(* Logix 5000 project; controller MV vendor 1 type 14 code 217 rev 31.11; software revision 31.00; part 21 of 53 *)
(* tags used below, declared in another part *)
   CheckTimeMask : INT;
   CWD : CHECKWORD_FLAGS;
   Delphi_Does_Eng_Func : BOOL;
   MC_CH2_DR1 : PlantItem;   // CH2_DR1
   MC_CH2_DR2 : PlantItem;   // CH2_DR2
   MC_CH2_DRAIN : PlantItem;   // CH2_DRAIN
   MC_CH2_DT1 : PlantItem;   // CH2_DT1
   MC_CH2_DT2 : PlantItem;   // CH2_DT2
   MC_CH2_LF1 : PlantItem;   // CH2_LF1
   MC_CH2_PR1 : PlantItem;   // CH2_PR1
   MC_CH2_R2R : PlantItem;   // CH2_R2R
   MC_CH2_R3R : PlantItem;   // CH2_R3R
   MC_CH2_R4R : PlantItem;   // CH2_R4R
   MC_CH2_R5R : PlantItem;   // CH2_R5R
   MC_CH2_R6R : PlantItem;   // CH2_R6R
   MC_CH2_RR : PlantItem;   // CH2_RR
   MC_N255 : INT[255];   // CHECKWORDS Plant item checkword s
   TempChecktime : DINT;
(* MC_Common, continued *)

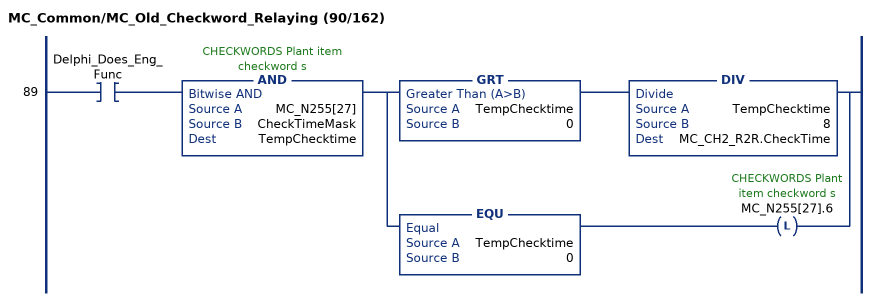
   [picture p361: MC_Common/MC_Old_Checkword_Relaying rungs 89-89]
   89: XIC(Delphi_Does_Eng_Func)AND(MC_N255[27],CheckTimeMask,TempChecktime)[GRT(TempChecktime,0) DIV(TempChecktime,8,MC_CH2_R2R.CheckTime) ,EQU(TempChecktime,0) OTL(MC_N255[27].6) ];
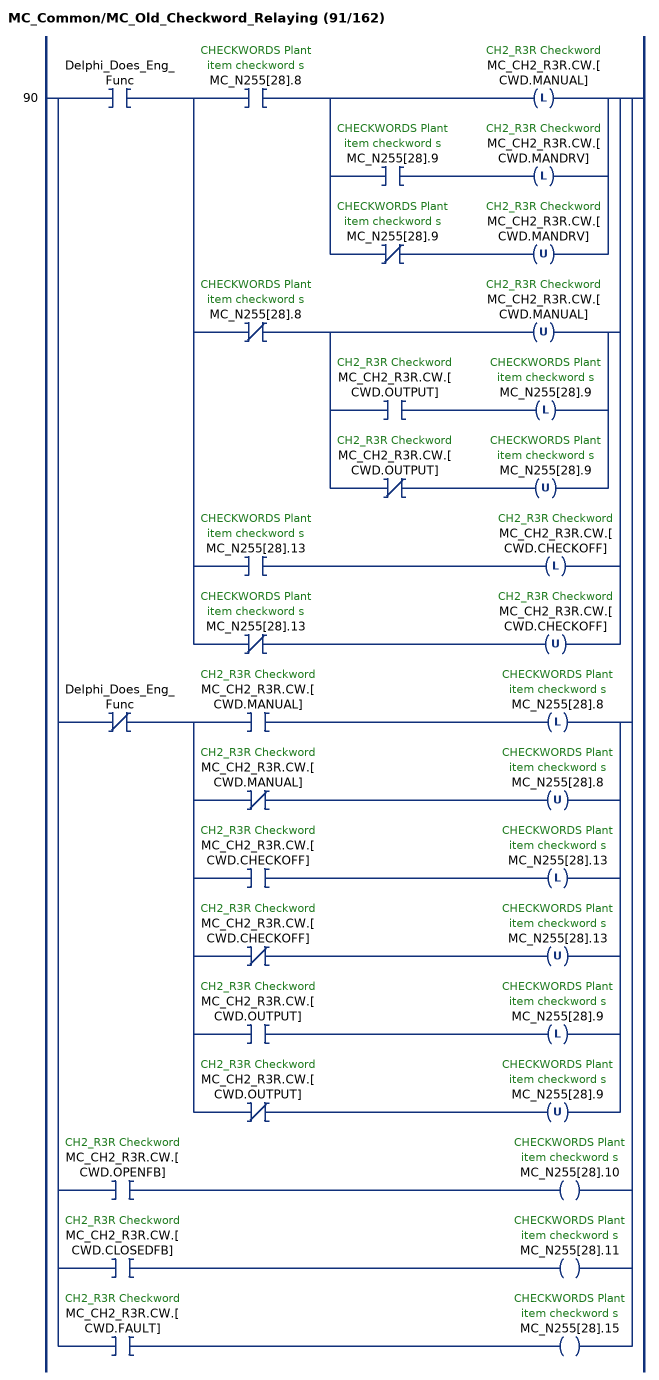
   90: [XIC(Delphi_Does_Eng_Func) [[XIC(MC_N255[28].8) [OTL(MC_CH2_R3R.CW.[CWD.MANUAL]) ,XIC(MC_N255[28].9) OTL(MC_CH2_R3R.CW.[CWD.MANDRV]) ,XIO(MC_N255[28].9) OTU(MC_CH2_R3R.CW.[CWD.MANDRV]) ] ,XIO(MC_N255[28].8) [OTU(MC_CH2_R3R.CW.[CWD.MANUAL]) ,[XIC(MC_CH2_R3R.CW.[CWD.OUTPUT]) OTL(MC_N255[28].9) ,XIO(MC_CH2_R3R.CW.[CWD.OUTPUT]) OTU(MC_N255[28].9) ] ] ] ,[XIC(MC_N255[28].13) OTL(MC_CH2_R3R.CW.[CWD.CHECKOFF]) ,XIO(MC_N255[28].13) OTU(MC_CH2_R3R.CW.[CWD.CHECKOFF]) ] ] ,XIO(Delphi_Does_Eng_Func) [[XIC(MC_CH2_R3R.CW.[CWD.MANUAL]) OTL(MC_N255[28].8) ,XIO(MC_CH2_R3R.CW.[CWD.MANUAL]) OTU(MC_N255[28].8) ] ,[XIC(MC_CH2_R3R.CW.[CWD.CHECKOFF]) OTL(MC_N255[28].13) ,XIO(MC_CH2_R3R.CW.[CWD.CHECKOFF]) OTU(MC_N255[28].13) ] ,[XIC(MC_CH2_R3R.CW.[CWD.OUTPUT]) OTL(MC_N255[28].9) ,XIO(MC_CH2_R3R.CW.[CWD.OUTPUT]) OTU(MC_N255[28].9) ] ] ,XIC(MC_CH2_R3R.CW.[CWD.OPENFB]) OTE(MC_N255[28].10) ,XIC(MC_CH2_R3R.CW.[CWD.CLOSEDFB]) OTE(MC_N255[28].11) ,XIC(MC_CH2_R3R.CW.[CWD.FAULT]) OTE(MC_N255[28].15) ];
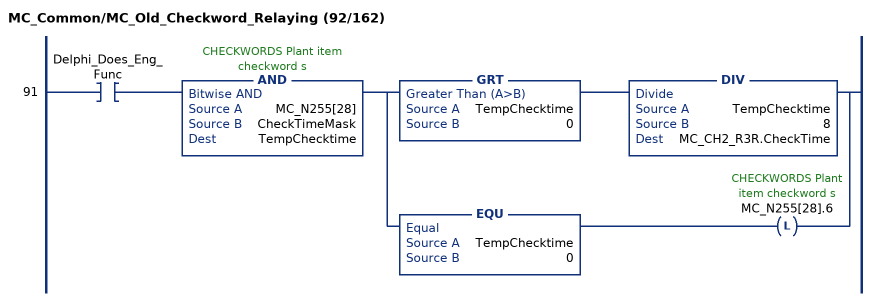
   91: XIC(Delphi_Does_Eng_Func)AND(MC_N255[28],CheckTimeMask,TempChecktime)[GRT(TempChecktime,0) DIV(TempChecktime,8,MC_CH2_R3R.CheckTime) ,EQU(TempChecktime,0) OTL(MC_N255[28].6) ];
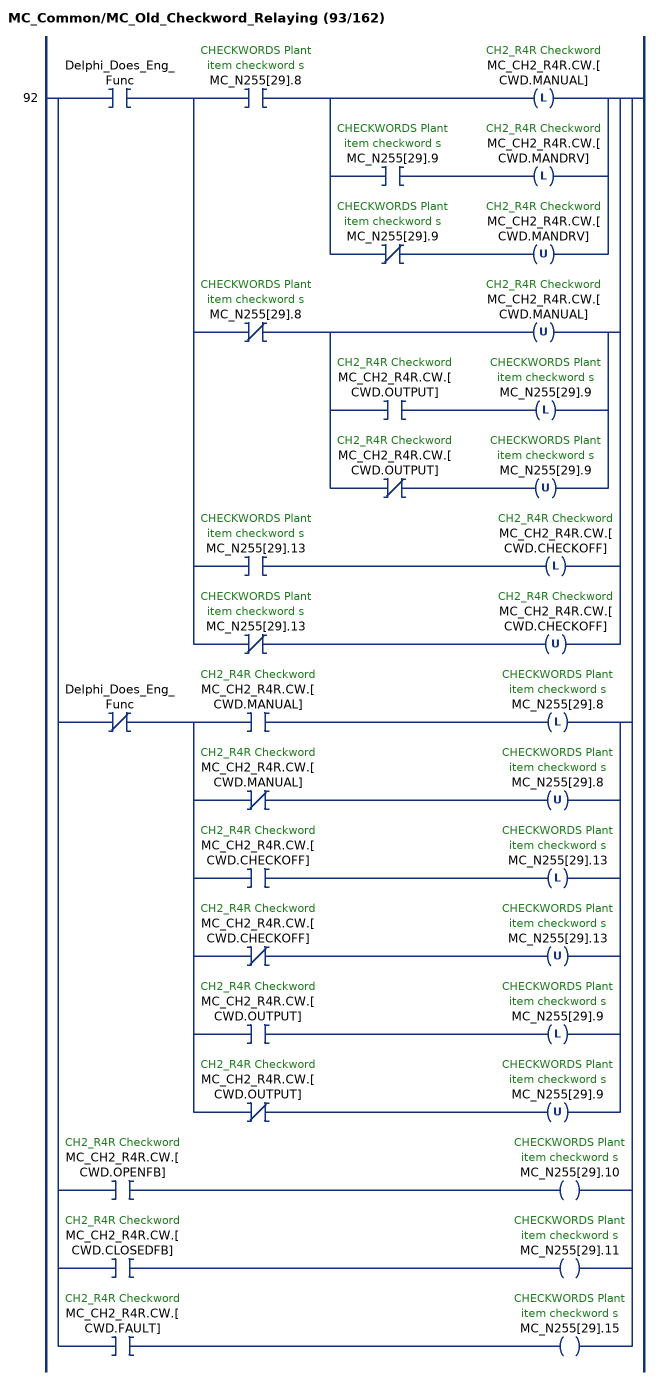
   92: [XIC(Delphi_Does_Eng_Func) [[XIC(MC_N255[29].8) [OTL(MC_CH2_R4R.CW.[CWD.MANUAL]) ,XIC(MC_N255[29].9) OTL(MC_CH2_R4R.CW.[CWD.MANDRV]) ,XIO(MC_N255[29].9) OTU(MC_CH2_R4R.CW.[CWD.MANDRV]) ] ,XIO(MC_N255[29].8) [OTU(MC_CH2_R4R.CW.[CWD.MANUAL]) ,[XIC(MC_CH2_R4R.CW.[CWD.OUTPUT]) OTL(MC_N255[29].9) ,XIO(MC_CH2_R4R.CW.[CWD.OUTPUT]) OTU(MC_N255[29].9) ] ] ] ,[XIC(MC_N255[29].13) OTL(MC_CH2_R4R.CW.[CWD.CHECKOFF]) ,XIO(MC_N255[29].13) OTU(MC_CH2_R4R.CW.[CWD.CHECKOFF]) ] ] ,XIO(Delphi_Does_Eng_Func) [[XIC(MC_CH2_R4R.CW.[CWD.MANUAL]) OTL(MC_N255[29].8) ,XIO(MC_CH2_R4R.CW.[CWD.MANUAL]) OTU(MC_N255[29].8) ] ,[XIC(MC_CH2_R4R.CW.[CWD.CHECKOFF]) OTL(MC_N255[29].13) ,XIO(MC_CH2_R4R.CW.[CWD.CHECKOFF]) OTU(MC_N255[29].13) ] ,[XIC(MC_CH2_R4R.CW.[CWD.OUTPUT]) OTL(MC_N255[29].9) ,XIO(MC_CH2_R4R.CW.[CWD.OUTPUT]) OTU(MC_N255[29].9) ] ] ,XIC(MC_CH2_R4R.CW.[CWD.OPENFB]) OTE(MC_N255[29].10) ,XIC(MC_CH2_R4R.CW.[CWD.CLOSEDFB]) OTE(MC_N255[29].11) ,XIC(MC_CH2_R4R.CW.[CWD.FAULT]) OTE(MC_N255[29].15) ];
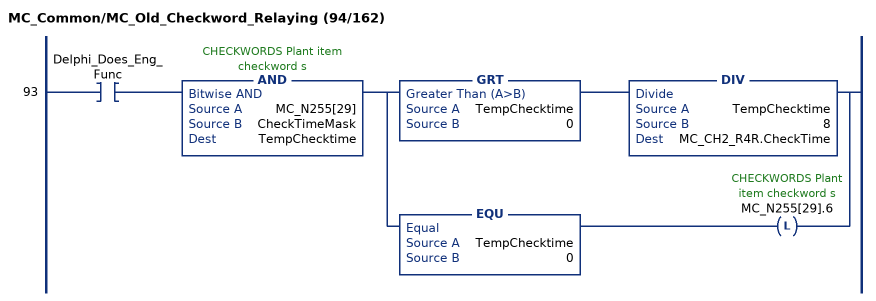
   93: XIC(Delphi_Does_Eng_Func)AND(MC_N255[29],CheckTimeMask,TempChecktime)[GRT(TempChecktime,0) DIV(TempChecktime,8,MC_CH2_R4R.CheckTime) ,EQU(TempChecktime,0) OTL(MC_N255[29].6) ];
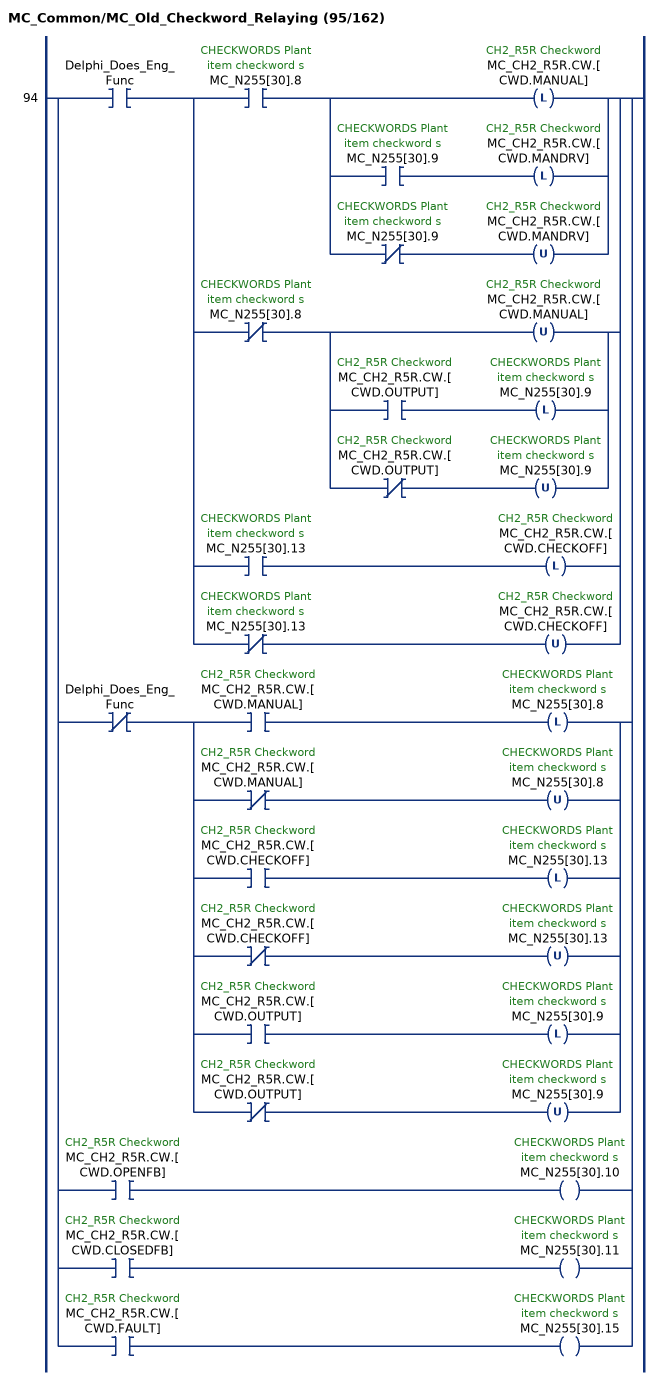
   94: [XIC(Delphi_Does_Eng_Func) [[XIC(MC_N255[30].8) [OTL(MC_CH2_R5R.CW.[CWD.MANUAL]) ,XIC(MC_N255[30].9) OTL(MC_CH2_R5R.CW.[CWD.MANDRV]) ,XIO(MC_N255[30].9) OTU(MC_CH2_R5R.CW.[CWD.MANDRV]) ] ,XIO(MC_N255[30].8) [OTU(MC_CH2_R5R.CW.[CWD.MANUAL]) ,[XIC(MC_CH2_R5R.CW.[CWD.OUTPUT]) OTL(MC_N255[30].9) ,XIO(MC_CH2_R5R.CW.[CWD.OUTPUT]) OTU(MC_N255[30].9) ] ] ] ,[XIC(MC_N255[30].13) OTL(MC_CH2_R5R.CW.[CWD.CHECKOFF]) ,XIO(MC_N255[30].13) OTU(MC_CH2_R5R.CW.[CWD.CHECKOFF]) ] ] ,XIO(Delphi_Does_Eng_Func) [[XIC(MC_CH2_R5R.CW.[CWD.MANUAL]) OTL(MC_N255[30].8) ,XIO(MC_CH2_R5R.CW.[CWD.MANUAL]) OTU(MC_N255[30].8) ] ,[XIC(MC_CH2_R5R.CW.[CWD.CHECKOFF]) OTL(MC_N255[30].13) ,XIO(MC_CH2_R5R.CW.[CWD.CHECKOFF]) OTU(MC_N255[30].13) ] ,[XIC(MC_CH2_R5R.CW.[CWD.OUTPUT]) OTL(MC_N255[30].9) ,XIO(MC_CH2_R5R.CW.[CWD.OUTPUT]) OTU(MC_N255[30].9) ] ] ,XIC(MC_CH2_R5R.CW.[CWD.OPENFB]) OTE(MC_N255[30].10) ,XIC(MC_CH2_R5R.CW.[CWD.CLOSEDFB]) OTE(MC_N255[30].11) ,XIC(MC_CH2_R5R.CW.[CWD.FAULT]) OTE(MC_N255[30].15) ];
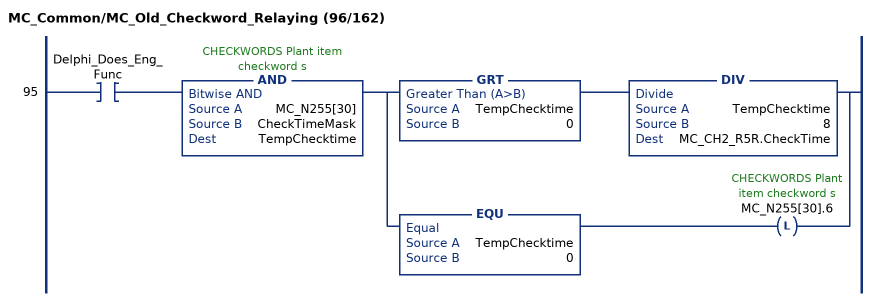
   95: XIC(Delphi_Does_Eng_Func)AND(MC_N255[30],CheckTimeMask,TempChecktime)[GRT(TempChecktime,0) DIV(TempChecktime,8,MC_CH2_R5R.CheckTime) ,EQU(TempChecktime,0) OTL(MC_N255[30].6) ];
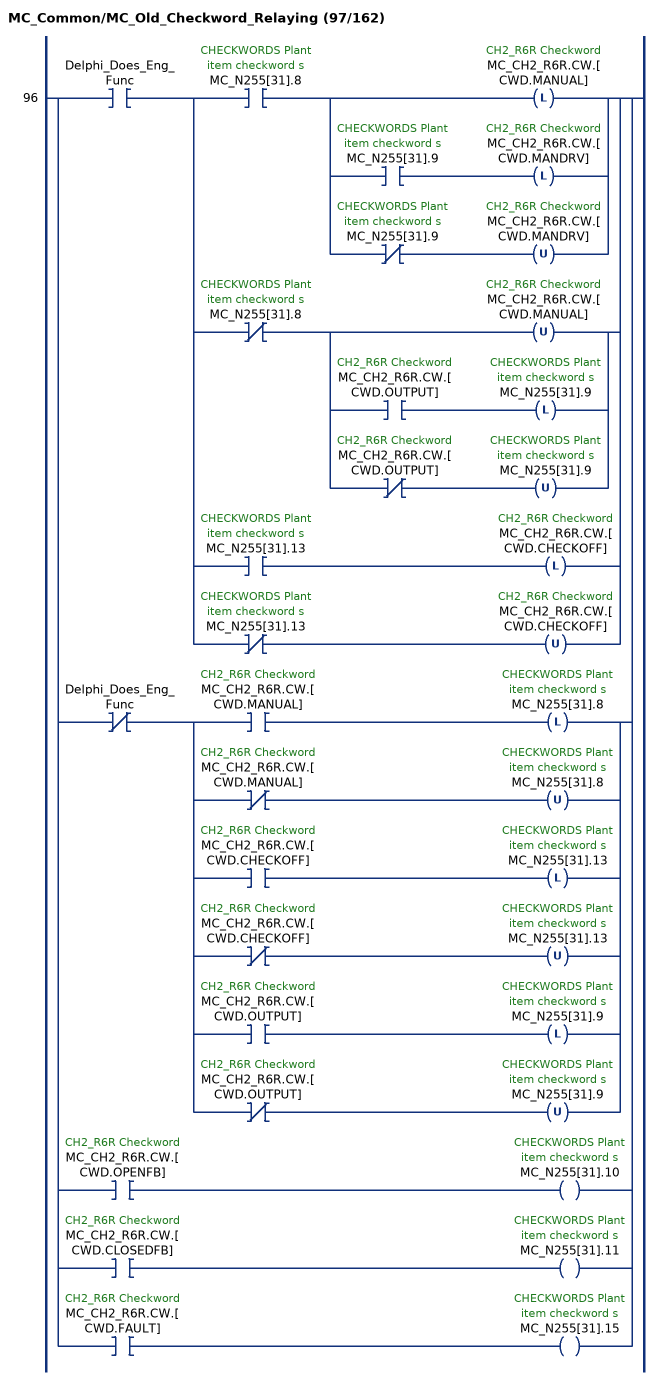
   96: [XIC(Delphi_Does_Eng_Func) [[XIC(MC_N255[31].8) [OTL(MC_CH2_R6R.CW.[CWD.MANUAL]) ,XIC(MC_N255[31].9) OTL(MC_CH2_R6R.CW.[CWD.MANDRV]) ,XIO(MC_N255[31].9) OTU(MC_CH2_R6R.CW.[CWD.MANDRV]) ] ,XIO(MC_N255[31].8) [OTU(MC_CH2_R6R.CW.[CWD.MANUAL]) ,[XIC(MC_CH2_R6R.CW.[CWD.OUTPUT]) OTL(MC_N255[31].9) ,XIO(MC_CH2_R6R.CW.[CWD.OUTPUT]) OTU(MC_N255[31].9) ] ] ] ,[XIC(MC_N255[31].13) OTL(MC_CH2_R6R.CW.[CWD.CHECKOFF]) ,XIO(MC_N255[31].13) OTU(MC_CH2_R6R.CW.[CWD.CHECKOFF]) ] ] ,XIO(Delphi_Does_Eng_Func) [[XIC(MC_CH2_R6R.CW.[CWD.MANUAL]) OTL(MC_N255[31].8) ,XIO(MC_CH2_R6R.CW.[CWD.MANUAL]) OTU(MC_N255[31].8) ] ,[XIC(MC_CH2_R6R.CW.[CWD.CHECKOFF]) OTL(MC_N255[31].13) ,XIO(MC_CH2_R6R.CW.[CWD.CHECKOFF]) OTU(MC_N255[31].13) ] ,[XIC(MC_CH2_R6R.CW.[CWD.OUTPUT]) OTL(MC_N255[31].9) ,XIO(MC_CH2_R6R.CW.[CWD.OUTPUT]) OTU(MC_N255[31].9) ] ] ,XIC(MC_CH2_R6R.CW.[CWD.OPENFB]) OTE(MC_N255[31].10) ,XIC(MC_CH2_R6R.CW.[CWD.CLOSEDFB]) OTE(MC_N255[31].11) ,XIC(MC_CH2_R6R.CW.[CWD.FAULT]) OTE(MC_N255[31].15) ];
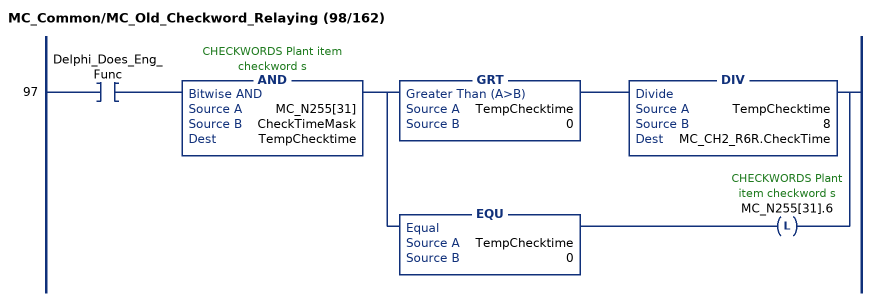
   97: XIC(Delphi_Does_Eng_Func)AND(MC_N255[31],CheckTimeMask,TempChecktime)[GRT(TempChecktime,0) DIV(TempChecktime,8,MC_CH2_R6R.CheckTime) ,EQU(TempChecktime,0) OTL(MC_N255[31].6) ];
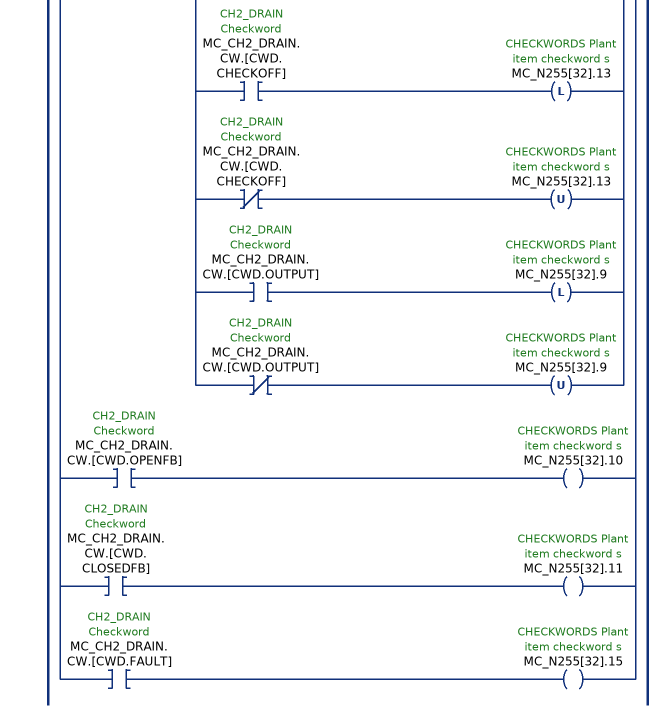
   98: [XIC(Delphi_Does_Eng_Func) [[XIC(MC_N255[32].8) [OTL(MC_CH2_DRAIN.CW.[CWD.MANUAL]) ,XIC(MC_N255[32].9) OTL(MC_CH2_DRAIN.CW.[CWD.MANDRV]) ,XIO(MC_N255[32].9) OTU(MC_CH2_DRAIN.CW.[CWD.MANDRV]) ] ,XIO(MC_N255[32].8) [OTU(MC_CH2_DRAIN.CW.[CWD.MANUAL]) ,[XIC(MC_CH2_DRAIN.CW.[CWD.OUTPUT]) OTL(MC_N255[32].9) ,XIO(MC_CH2_DRAIN.CW.[CWD.OUTPUT]) OTU(MC_N255[32].9) ] ] ] ,[XIC(MC_N255[32].13) OTL(MC_CH2_DRAIN.CW.[CWD.CHECKOFF]) ,XIO(MC_N255[32].13) OTU(MC_CH2_DRAIN.CW.[CWD.CHECKOFF]) ] ] ,XIO(Delphi_Does_Eng_Func) [[XIC(MC_CH2_DRAIN.CW.[CWD.MANUAL]) OTL(MC_N255[32].8) ,XIO(MC_CH2_DRAIN.CW.[CWD.MANUAL]) OTU(MC_N255[32].8) ] ,[XIC(MC_CH2_DRAIN.CW.[CWD.CHECKOFF]) OTL(MC_N255[32].13) ,XIO(MC_CH2_DRAIN.CW.[CWD.CHECKOFF]) OTU(MC_N255[32].13) ] ,[XIC(MC_CH2_DRAIN.CW.[CWD.OUTPUT]) OTL(MC_N255[32].9) ,XIO(MC_CH2_DRAIN.CW.[CWD.OUTPUT]) OTU(MC_N255[32].9) ] ] ,XIC(MC_CH2_DRAIN.CW.[CWD.OPENFB]) OTE(MC_N255[32].10) ,XIC(MC_CH2_DRAIN.CW.[CWD.CLOSEDFB]) OTE(MC_N255[32].11) ,XIC(MC_CH2_DRAIN.CW.[CWD.FAULT]) OTE(MC_N255[32].15) ];
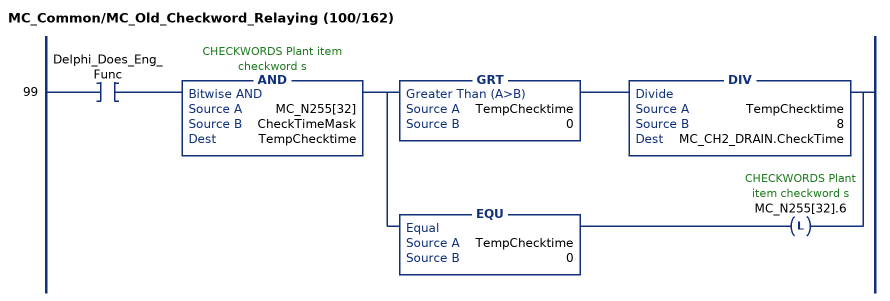
   99: XIC(Delphi_Does_Eng_Func)AND(MC_N255[32],CheckTimeMask,TempChecktime)[GRT(TempChecktime,0) DIV(TempChecktime,8,MC_CH2_DRAIN.CheckTime) ,EQU(TempChecktime,0) OTL(MC_N255[32].6) ];
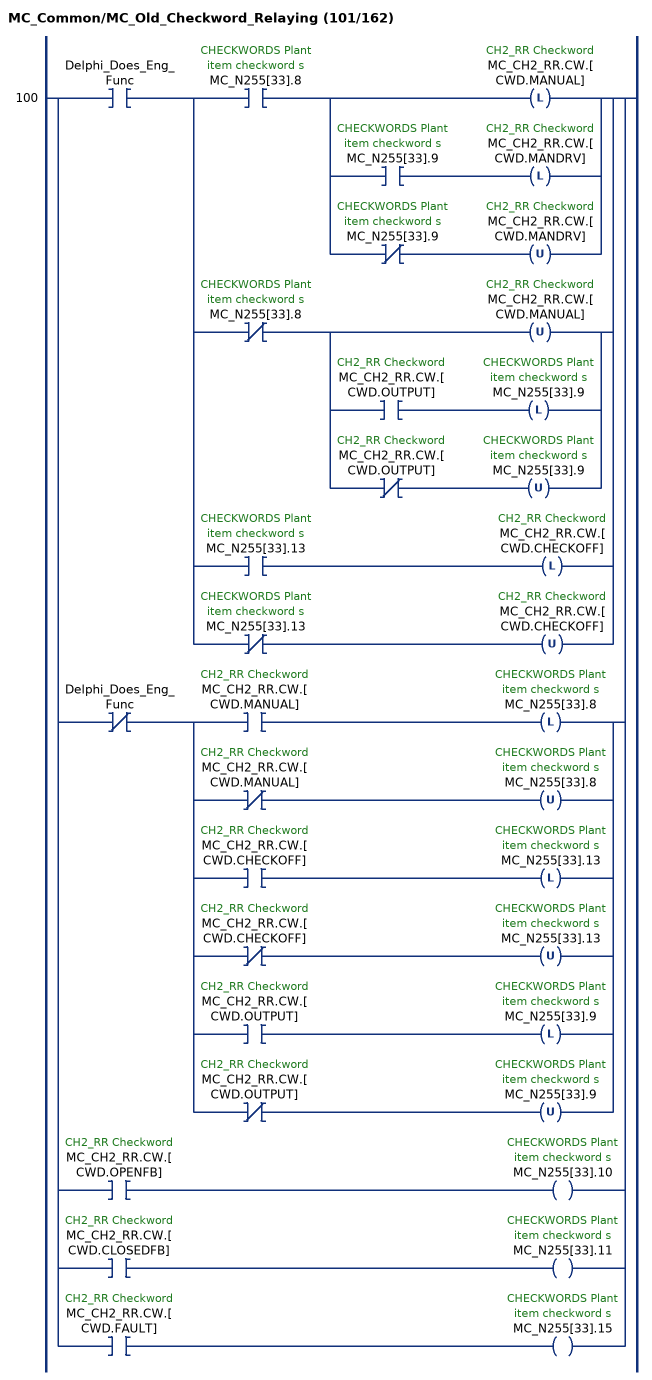
   100: [XIC(Delphi_Does_Eng_Func) [[XIC(MC_N255[33].8) [OTL(MC_CH2_RR.CW.[CWD.MANUAL]) ,XIC(MC_N255[33].9) OTL(MC_CH2_RR.CW.[CWD.MANDRV]) ,XIO(MC_N255[33].9) OTU(MC_CH2_RR.CW.[CWD.MANDRV]) ] ,XIO(MC_N255[33].8) [OTU(MC_CH2_RR.CW.[CWD.MANUAL]) ,[XIC(MC_CH2_RR.CW.[CWD.OUTPUT]) OTL(MC_N255[33].9) ,XIO(MC_CH2_RR.CW.[CWD.OUTPUT]) OTU(MC_N255[33].9) ] ] ] ,[XIC(MC_N255[33].13) OTL(MC_CH2_RR.CW.[CWD.CHECKOFF]) ,XIO(MC_N255[33].13) OTU(MC_CH2_RR.CW.[CWD.CHECKOFF]) ] ] ,XIO(Delphi_Does_Eng_Func) [[XIC(MC_CH2_RR.CW.[CWD.MANUAL]) OTL(MC_N255[33].8) ,XIO(MC_CH2_RR.CW.[CWD.MANUAL]) OTU(MC_N255[33].8) ] ,[XIC(MC_CH2_RR.CW.[CWD.CHECKOFF]) OTL(MC_N255[33].13) ,XIO(MC_CH2_RR.CW.[CWD.CHECKOFF]) OTU(MC_N255[33].13) ] ,[XIC(MC_CH2_RR.CW.[CWD.OUTPUT]) OTL(MC_N255[33].9) ,XIO(MC_CH2_RR.CW.[CWD.OUTPUT]) OTU(MC_N255[33].9) ] ] ,XIC(MC_CH2_RR.CW.[CWD.OPENFB]) OTE(MC_N255[33].10) ,XIC(MC_CH2_RR.CW.[CWD.CLOSEDFB]) OTE(MC_N255[33].11) ,XIC(MC_CH2_RR.CW.[CWD.FAULT]) OTE(MC_N255[33].15) ];
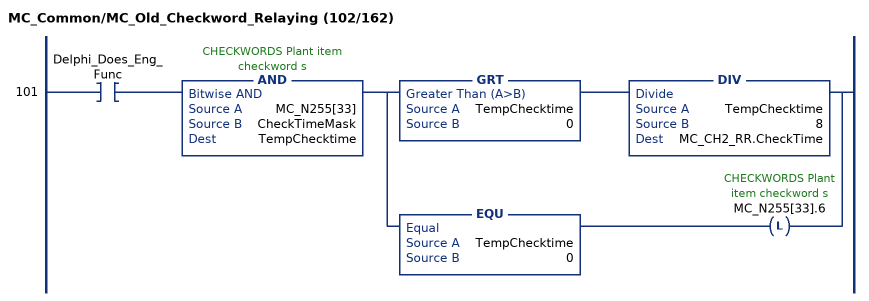
   101: XIC(Delphi_Does_Eng_Func)AND(MC_N255[33],CheckTimeMask,TempChecktime)[GRT(TempChecktime,0) DIV(TempChecktime,8,MC_CH2_RR.CheckTime) ,EQU(TempChecktime,0) OTL(MC_N255[33].6) ];
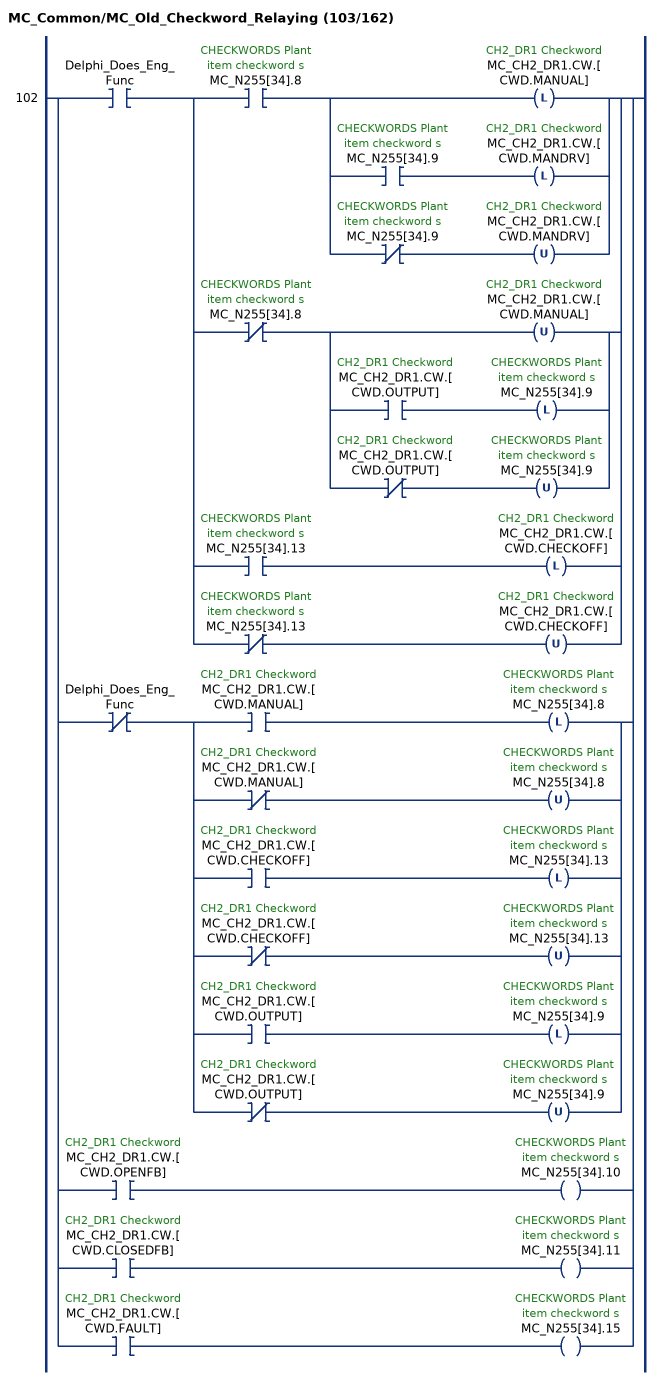
   102: [XIC(Delphi_Does_Eng_Func) [[XIC(MC_N255[34].8) [OTL(MC_CH2_DR1.CW.[CWD.MANUAL]) ,XIC(MC_N255[34].9) OTL(MC_CH2_DR1.CW.[CWD.MANDRV]) ,XIO(MC_N255[34].9) OTU(MC_CH2_DR1.CW.[CWD.MANDRV]) ] ,XIO(MC_N255[34].8) [OTU(MC_CH2_DR1.CW.[CWD.MANUAL]) ,[XIC(MC_CH2_DR1.CW.[CWD.OUTPUT]) OTL(MC_N255[34].9) ,XIO(MC_CH2_DR1.CW.[CWD.OUTPUT]) OTU(MC_N255[34].9) ] ] ] ,[XIC(MC_N255[34].13) OTL(MC_CH2_DR1.CW.[CWD.CHECKOFF]) ,XIO(MC_N255[34].13) OTU(MC_CH2_DR1.CW.[CWD.CHECKOFF]) ] ] ,XIO(Delphi_Does_Eng_Func) [[XIC(MC_CH2_DR1.CW.[CWD.MANUAL]) OTL(MC_N255[34].8) ,XIO(MC_CH2_DR1.CW.[CWD.MANUAL]) OTU(MC_N255[34].8) ] ,[XIC(MC_CH2_DR1.CW.[CWD.CHECKOFF]) OTL(MC_N255[34].13) ,XIO(MC_CH2_DR1.CW.[CWD.CHECKOFF]) OTU(MC_N255[34].13) ] ,[XIC(MC_CH2_DR1.CW.[CWD.OUTPUT]) OTL(MC_N255[34].9) ,XIO(MC_CH2_DR1.CW.[CWD.OUTPUT]) OTU(MC_N255[34].9) ] ] ,XIC(MC_CH2_DR1.CW.[CWD.OPENFB]) OTE(MC_N255[34].10) ,XIC(MC_CH2_DR1.CW.[CWD.CLOSEDFB]) OTE(MC_N255[34].11) ,XIC(MC_CH2_DR1.CW.[CWD.FAULT]) OTE(MC_N255[34].15) ];
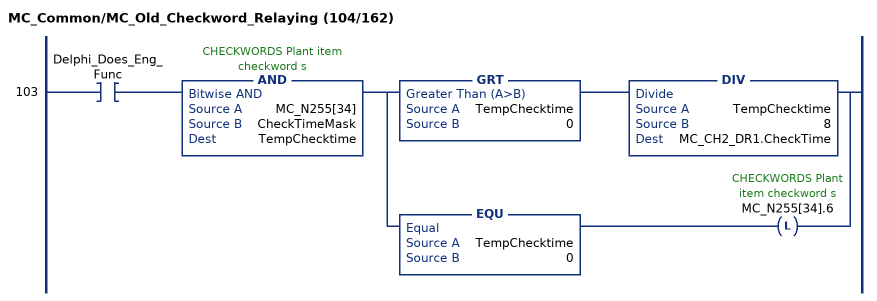
   103: XIC(Delphi_Does_Eng_Func)AND(MC_N255[34],CheckTimeMask,TempChecktime)[GRT(TempChecktime,0) DIV(TempChecktime,8,MC_CH2_DR1.CheckTime) ,EQU(TempChecktime,0) OTL(MC_N255[34].6) ];
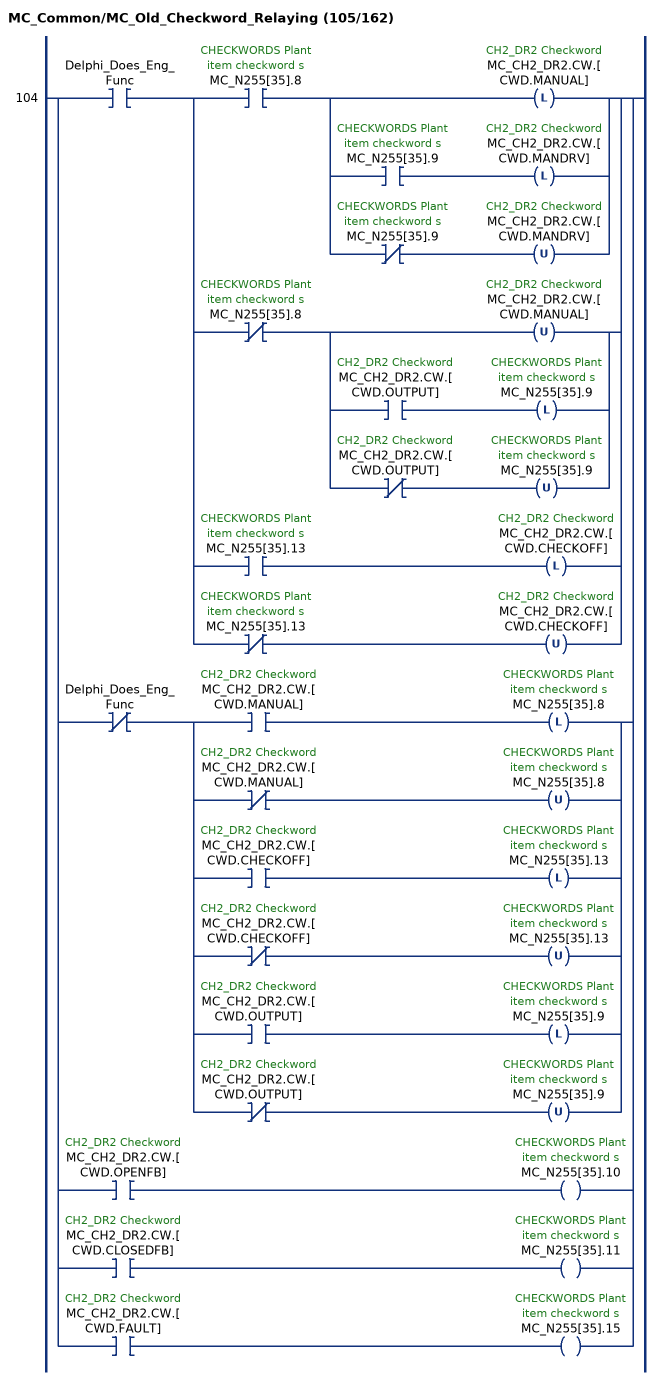
   104: [XIC(Delphi_Does_Eng_Func) [[XIC(MC_N255[35].8) [OTL(MC_CH2_DR2.CW.[CWD.MANUAL]) ,XIC(MC_N255[35].9) OTL(MC_CH2_DR2.CW.[CWD.MANDRV]) ,XIO(MC_N255[35].9) OTU(MC_CH2_DR2.CW.[CWD.MANDRV]) ] ,XIO(MC_N255[35].8) [OTU(MC_CH2_DR2.CW.[CWD.MANUAL]) ,[XIC(MC_CH2_DR2.CW.[CWD.OUTPUT]) OTL(MC_N255[35].9) ,XIO(MC_CH2_DR2.CW.[CWD.OUTPUT]) OTU(MC_N255[35].9) ] ] ] ,[XIC(MC_N255[35].13) OTL(MC_CH2_DR2.CW.[CWD.CHECKOFF]) ,XIO(MC_N255[35].13) OTU(MC_CH2_DR2.CW.[CWD.CHECKOFF]) ] ] ,XIO(Delphi_Does_Eng_Func) [[XIC(MC_CH2_DR2.CW.[CWD.MANUAL]) OTL(MC_N255[35].8) ,XIO(MC_CH2_DR2.CW.[CWD.MANUAL]) OTU(MC_N255[35].8) ] ,[XIC(MC_CH2_DR2.CW.[CWD.CHECKOFF]) OTL(MC_N255[35].13) ,XIO(MC_CH2_DR2.CW.[CWD.CHECKOFF]) OTU(MC_N255[35].13) ] ,[XIC(MC_CH2_DR2.CW.[CWD.OUTPUT]) OTL(MC_N255[35].9) ,XIO(MC_CH2_DR2.CW.[CWD.OUTPUT]) OTU(MC_N255[35].9) ] ] ,XIC(MC_CH2_DR2.CW.[CWD.OPENFB]) OTE(MC_N255[35].10) ,XIC(MC_CH2_DR2.CW.[CWD.CLOSEDFB]) OTE(MC_N255[35].11) ,XIC(MC_CH2_DR2.CW.[CWD.FAULT]) OTE(MC_N255[35].15) ];
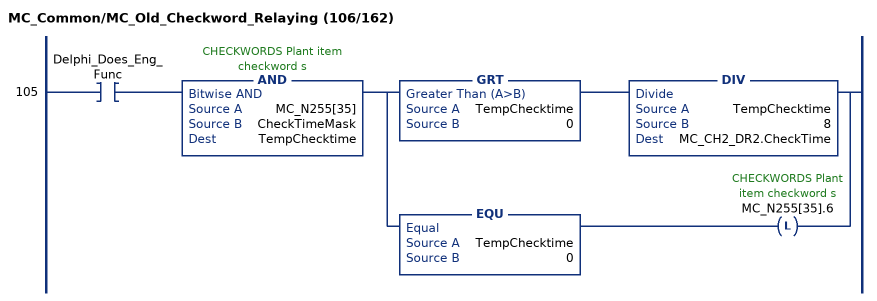
   105: XIC(Delphi_Does_Eng_Func)AND(MC_N255[35],CheckTimeMask,TempChecktime)[GRT(TempChecktime,0) DIV(TempChecktime,8,MC_CH2_DR2.CheckTime) ,EQU(TempChecktime,0) OTL(MC_N255[35].6) ];
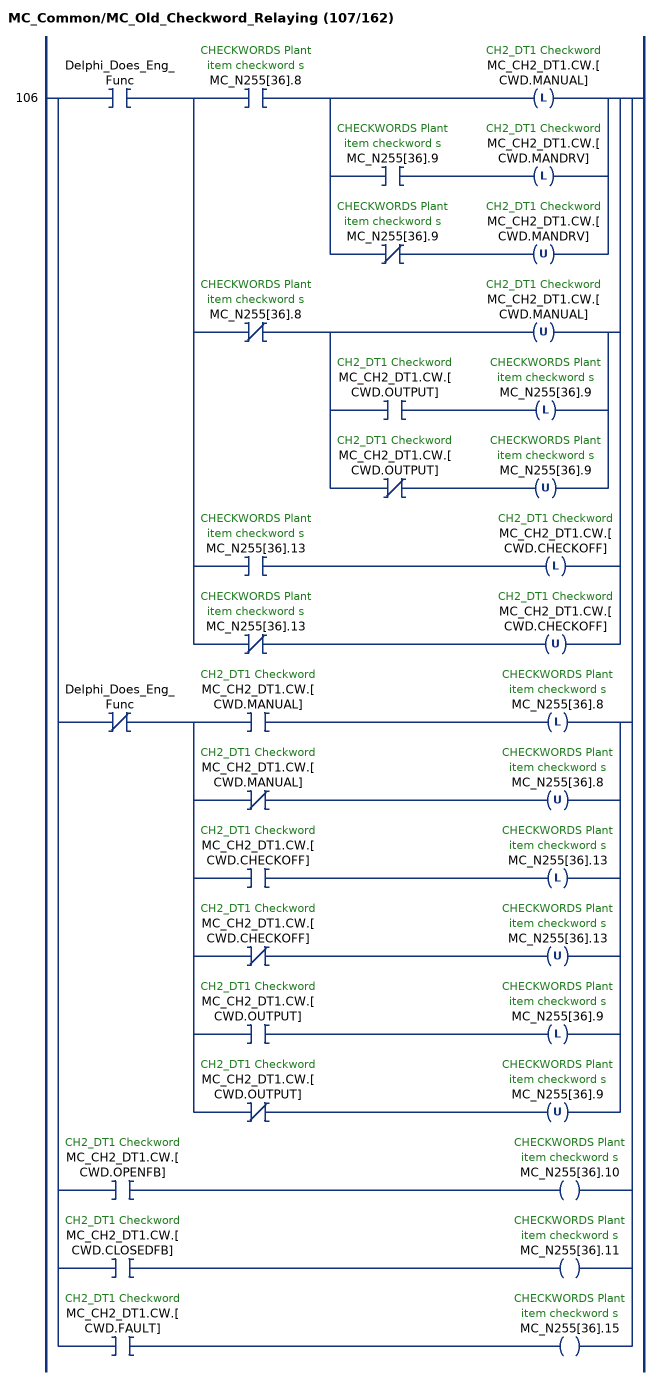
   106: [XIC(Delphi_Does_Eng_Func) [[XIC(MC_N255[36].8) [OTL(MC_CH2_DT1.CW.[CWD.MANUAL]) ,XIC(MC_N255[36].9) OTL(MC_CH2_DT1.CW.[CWD.MANDRV]) ,XIO(MC_N255[36].9) OTU(MC_CH2_DT1.CW.[CWD.MANDRV]) ] ,XIO(MC_N255[36].8) [OTU(MC_CH2_DT1.CW.[CWD.MANUAL]) ,[XIC(MC_CH2_DT1.CW.[CWD.OUTPUT]) OTL(MC_N255[36].9) ,XIO(MC_CH2_DT1.CW.[CWD.OUTPUT]) OTU(MC_N255[36].9) ] ] ] ,[XIC(MC_N255[36].13) OTL(MC_CH2_DT1.CW.[CWD.CHECKOFF]) ,XIO(MC_N255[36].13) OTU(MC_CH2_DT1.CW.[CWD.CHECKOFF]) ] ] ,XIO(Delphi_Does_Eng_Func) [[XIC(MC_CH2_DT1.CW.[CWD.MANUAL]) OTL(MC_N255[36].8) ,XIO(MC_CH2_DT1.CW.[CWD.MANUAL]) OTU(MC_N255[36].8) ] ,[XIC(MC_CH2_DT1.CW.[CWD.CHECKOFF]) OTL(MC_N255[36].13) ,XIO(MC_CH2_DT1.CW.[CWD.CHECKOFF]) OTU(MC_N255[36].13) ] ,[XIC(MC_CH2_DT1.CW.[CWD.OUTPUT]) OTL(MC_N255[36].9) ,XIO(MC_CH2_DT1.CW.[CWD.OUTPUT]) OTU(MC_N255[36].9) ] ] ,XIC(MC_CH2_DT1.CW.[CWD.OPENFB]) OTE(MC_N255[36].10) ,XIC(MC_CH2_DT1.CW.[CWD.CLOSEDFB]) OTE(MC_N255[36].11) ,XIC(MC_CH2_DT1.CW.[CWD.FAULT]) OTE(MC_N255[36].15) ];
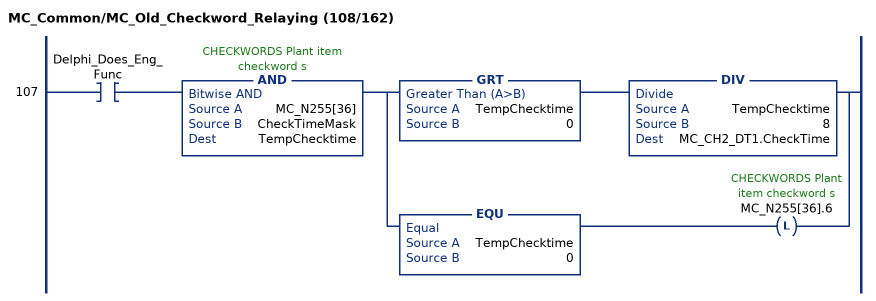
   107: XIC(Delphi_Does_Eng_Func)AND(MC_N255[36],CheckTimeMask,TempChecktime)[GRT(TempChecktime,0) DIV(TempChecktime,8,MC_CH2_DT1.CheckTime) ,EQU(TempChecktime,0) OTL(MC_N255[36].6) ];
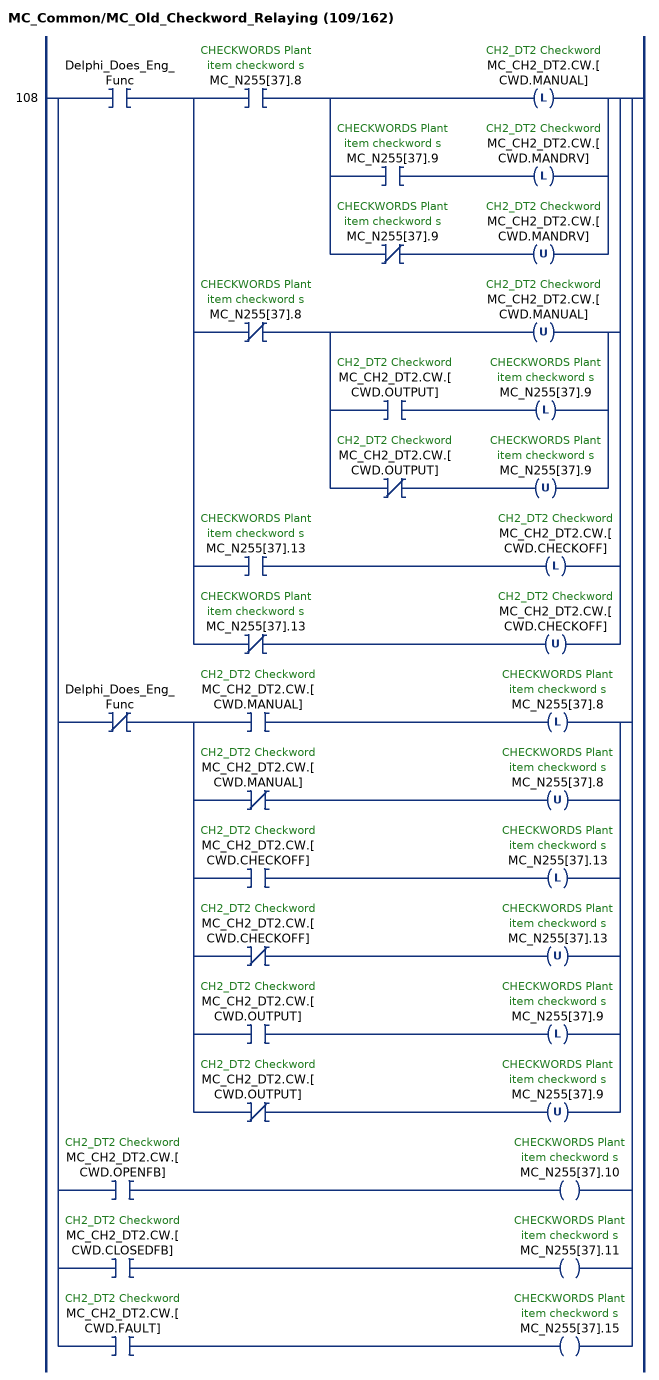
   108: [XIC(Delphi_Does_Eng_Func) [[XIC(MC_N255[37].8) [OTL(MC_CH2_DT2.CW.[CWD.MANUAL]) ,XIC(MC_N255[37].9) OTL(MC_CH2_DT2.CW.[CWD.MANDRV]) ,XIO(MC_N255[37].9) OTU(MC_CH2_DT2.CW.[CWD.MANDRV]) ] ,XIO(MC_N255[37].8) [OTU(MC_CH2_DT2.CW.[CWD.MANUAL]) ,[XIC(MC_CH2_DT2.CW.[CWD.OUTPUT]) OTL(MC_N255[37].9) ,XIO(MC_CH2_DT2.CW.[CWD.OUTPUT]) OTU(MC_N255[37].9) ] ] ] ,[XIC(MC_N255[37].13) OTL(MC_CH2_DT2.CW.[CWD.CHECKOFF]) ,XIO(MC_N255[37].13) OTU(MC_CH2_DT2.CW.[CWD.CHECKOFF]) ] ] ,XIO(Delphi_Does_Eng_Func) [[XIC(MC_CH2_DT2.CW.[CWD.MANUAL]) OTL(MC_N255[37].8) ,XIO(MC_CH2_DT2.CW.[CWD.MANUAL]) OTU(MC_N255[37].8) ] ,[XIC(MC_CH2_DT2.CW.[CWD.CHECKOFF]) OTL(MC_N255[37].13) ,XIO(MC_CH2_DT2.CW.[CWD.CHECKOFF]) OTU(MC_N255[37].13) ] ,[XIC(MC_CH2_DT2.CW.[CWD.OUTPUT]) OTL(MC_N255[37].9) ,XIO(MC_CH2_DT2.CW.[CWD.OUTPUT]) OTU(MC_N255[37].9) ] ] ,XIC(MC_CH2_DT2.CW.[CWD.OPENFB]) OTE(MC_N255[37].10) ,XIC(MC_CH2_DT2.CW.[CWD.CLOSEDFB]) OTE(MC_N255[37].11) ,XIC(MC_CH2_DT2.CW.[CWD.FAULT]) OTE(MC_N255[37].15) ];
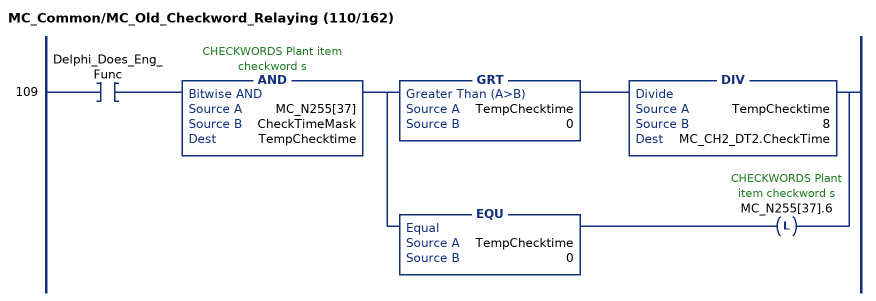
   109: XIC(Delphi_Does_Eng_Func)AND(MC_N255[37],CheckTimeMask,TempChecktime)[GRT(TempChecktime,0) DIV(TempChecktime,8,MC_CH2_DT2.CheckTime) ,EQU(TempChecktime,0) OTL(MC_N255[37].6) ];
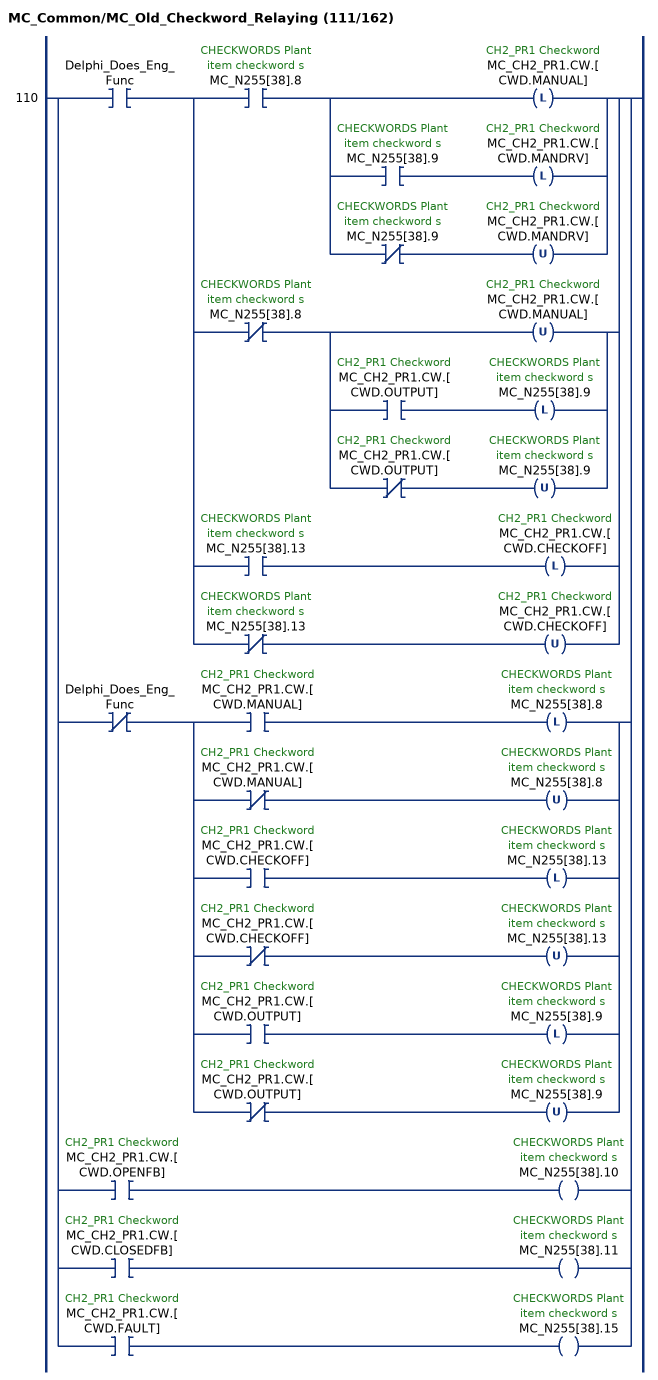
   110: [XIC(Delphi_Does_Eng_Func) [[XIC(MC_N255[38].8) [OTL(MC_CH2_PR1.CW.[CWD.MANUAL]) ,XIC(MC_N255[38].9) OTL(MC_CH2_PR1.CW.[CWD.MANDRV]) ,XIO(MC_N255[38].9) OTU(MC_CH2_PR1.CW.[CWD.MANDRV]) ] ,XIO(MC_N255[38].8) [OTU(MC_CH2_PR1.CW.[CWD.MANUAL]) ,[XIC(MC_CH2_PR1.CW.[CWD.OUTPUT]) OTL(MC_N255[38].9) ,XIO(MC_CH2_PR1.CW.[CWD.OUTPUT]) OTU(MC_N255[38].9) ] ] ] ,[XIC(MC_N255[38].13) OTL(MC_CH2_PR1.CW.[CWD.CHECKOFF]) ,XIO(MC_N255[38].13) OTU(MC_CH2_PR1.CW.[CWD.CHECKOFF]) ] ] ,XIO(Delphi_Does_Eng_Func) [[XIC(MC_CH2_PR1.CW.[CWD.MANUAL]) OTL(MC_N255[38].8) ,XIO(MC_CH2_PR1.CW.[CWD.MANUAL]) OTU(MC_N255[38].8) ] ,[XIC(MC_CH2_PR1.CW.[CWD.CHECKOFF]) OTL(MC_N255[38].13) ,XIO(MC_CH2_PR1.CW.[CWD.CHECKOFF]) OTU(MC_N255[38].13) ] ,[XIC(MC_CH2_PR1.CW.[CWD.OUTPUT]) OTL(MC_N255[38].9) ,XIO(MC_CH2_PR1.CW.[CWD.OUTPUT]) OTU(MC_N255[38].9) ] ] ,XIC(MC_CH2_PR1.CW.[CWD.OPENFB]) OTE(MC_N255[38].10) ,XIC(MC_CH2_PR1.CW.[CWD.CLOSEDFB]) OTE(MC_N255[38].11) ,XIC(MC_CH2_PR1.CW.[CWD.FAULT]) OTE(MC_N255[38].15) ];
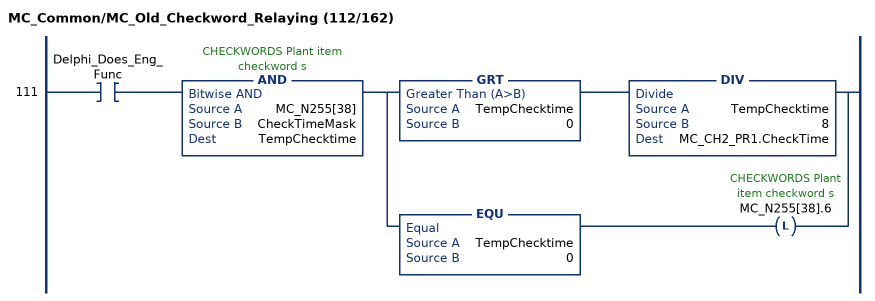
   111: XIC(Delphi_Does_Eng_Func)AND(MC_N255[38],CheckTimeMask,TempChecktime)[GRT(TempChecktime,0) DIV(TempChecktime,8,MC_CH2_PR1.CheckTime) ,EQU(TempChecktime,0) OTL(MC_N255[38].6) ];
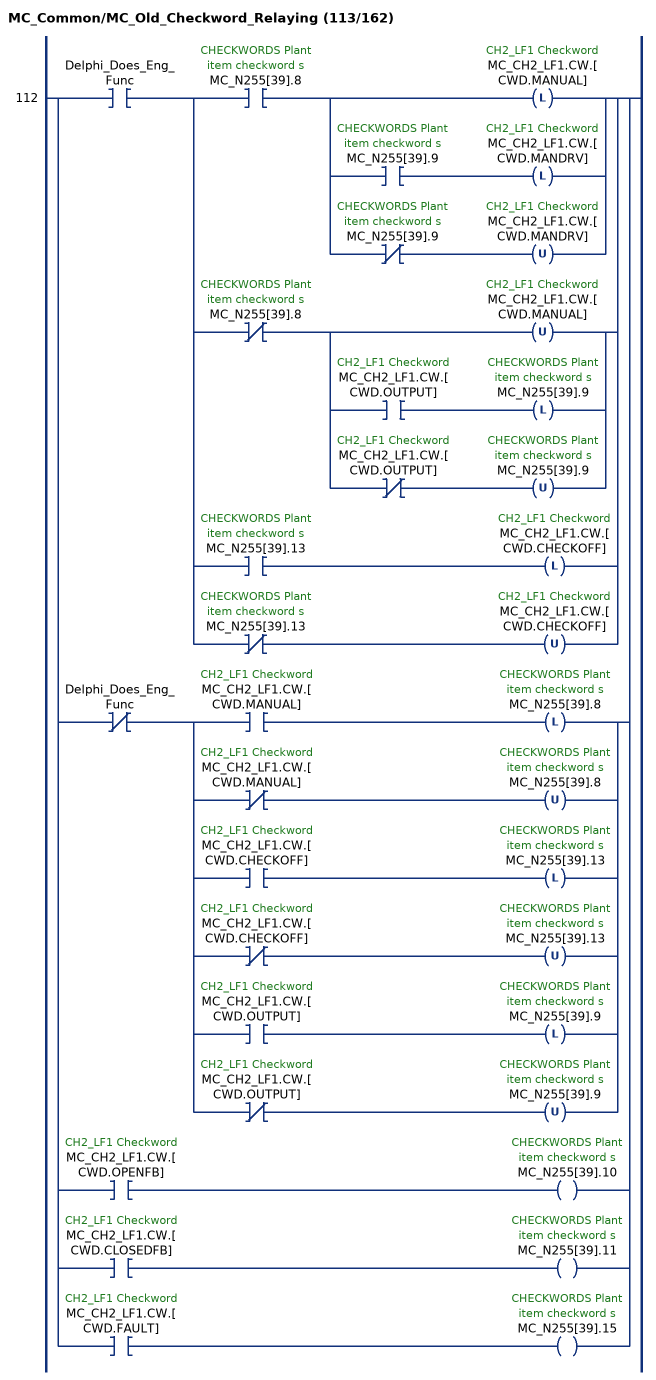
   112: [XIC(Delphi_Does_Eng_Func) [[XIC(MC_N255[39].8) [OTL(MC_CH2_LF1.CW.[CWD.MANUAL]) ,XIC(MC_N255[39].9) OTL(MC_CH2_LF1.CW.[CWD.MANDRV]) ,XIO(MC_N255[39].9) OTU(MC_CH2_LF1.CW.[CWD.MANDRV]) ] ,XIO(MC_N255[39].8) [OTU(MC_CH2_LF1.CW.[CWD.MANUAL]) ,[XIC(MC_CH2_LF1.CW.[CWD.OUTPUT]) OTL(MC_N255[39].9) ,XIO(MC_CH2_LF1.CW.[CWD.OUTPUT]) OTU(MC_N255[39].9) ] ] ] ,[XIC(MC_N255[39].13) OTL(MC_CH2_LF1.CW.[CWD.CHECKOFF]) ,XIO(MC_N255[39].13) OTU(MC_CH2_LF1.CW.[CWD.CHECKOFF]) ] ] ,XIO(Delphi_Does_Eng_Func) [[XIC(MC_CH2_LF1.CW.[CWD.MANUAL]) OTL(MC_N255[39].8) ,XIO(MC_CH2_LF1.CW.[CWD.MANUAL]) OTU(MC_N255[39].8) ] ,[XIC(MC_CH2_LF1.CW.[CWD.CHECKOFF]) OTL(MC_N255[39].13) ,XIO(MC_CH2_LF1.CW.[CWD.CHECKOFF]) OTU(MC_N255[39].13) ] ,[XIC(MC_CH2_LF1.CW.[CWD.OUTPUT]) OTL(MC_N255[39].9) ,XIO(MC_CH2_LF1.CW.[CWD.OUTPUT]) OTU(MC_N255[39].9) ] ] ,XIC(MC_CH2_LF1.CW.[CWD.OPENFB]) OTE(MC_N255[39].10) ,XIC(MC_CH2_LF1.CW.[CWD.CLOSEDFB]) OTE(MC_N255[39].11) ,XIC(MC_CH2_LF1.CW.[CWD.FAULT]) OTE(MC_N255[39].15) ];
